   	OWF_Key[436,9]:=1170757502;
   	OWF_Key[436,10]:=379063934;
   	OWF_Key[436,11]:=939425324;
   	OWF_Key[436,12]:=1571077433;
   	OWF_Key[436,13]:=386926956;
   	OWF_Key[436,14]:=1253683460;
   	OWF_Key[436,15]:=1978140769;
   	OWF_Key[436,16]:=969971513;
   	OWF_Key[437,0]:=1843141582;
   	OWF_Key[437,1]:=1139180362;
   	OWF_Key[437,2]:=1967511731;
   	OWF_Key[437,3]:=1290649002;
   	OWF_Key[437,4]:=1378760868;
   	OWF_Key[437,5]:=1424739908;
   	OWF_Key[437,6]:=88097231;
   	OWF_Key[437,7]:=835055186;
   	OWF_Key[437,8]:=1627536833;
   	OWF_Key[437,9]:=543176006;
   	OWF_Key[437,10]:=1462679088;
   	OWF_Key[437,11]:=893832072;
   	OWF_Key[437,12]:=149893027;
   	OWF_Key[437,13]:=919941861;
   	OWF_Key[437,14]:=1244070675;
   	OWF_Key[437,15]:=720720483;
   	OWF_Key[437,16]:=106207793;
   	OWF_Key[438,0]:=1266683906;
   	OWF_Key[438,1]:=1923048867;
   	OWF_Key[438,2]:=1845235682;
   	OWF_Key[438,3]:=1052576015;
   	OWF_Key[438,4]:=621819626;
   	OWF_Key[438,5]:=249692926;
   	OWF_Key[438,6]:=969832967;
   	OWF_Key[438,7]:=766223670;
   	OWF_Key[438,8]:=1411344155;
   	OWF_Key[438,9]:=1650208802;
   	OWF_Key[438,10]:=103954679;
   	OWF_Key[438,11]:=1231682890;
   	OWF_Key[438,12]:=1324790258;
   	OWF_Key[438,13]:=615786523;
   	OWF_Key[438,14]:=414858455;
   	OWF_Key[438,15]:=939305588;
   	OWF_Key[438,16]:=719104723;
   	OWF_Key[439,0]:=1992499359;
   	OWF_Key[439,1]:=251323729;
   	OWF_Key[439,2]:=600659015;
   	OWF_Key[439,3]:=1403077275;
   	OWF_Key[439,4]:=628364857;
   	OWF_Key[439,5]:=1823764687;
   	OWF_Key[439,6]:=631857018;
   	OWF_Key[439,7]:=1931716673;
   	OWF_Key[439,8]:=428827108;
   	OWF_Key[439,9]:=1029064288;
   	OWF_Key[439,10]:=1492699981;
   	OWF_Key[439,11]:=611446466;
   	OWF_Key[439,12]:=289686517;
   	OWF_Key[439,13]:=1524542361;
   	OWF_Key[439,14]:=69099460;
   	OWF_Key[439,15]:=1294673003;
   	OWF_Key[439,16]:=2029874974;
   	OWF_Key[440,0]:=267240957;
   	OWF_Key[440,1]:=1397447859;
   	OWF_Key[440,2]:=766044100;
   	OWF_Key[440,3]:=1128726900;
   	OWF_Key[440,4]:=808363166;
   	OWF_Key[440,5]:=1558535267;
   	OWF_Key[440,6]:=1447582414;
   	OWF_Key[440,7]:=964974356;
   	OWF_Key[440,8]:=1784322886;
   	OWF_Key[440,9]:=443035495;
   	OWF_Key[440,10]:=820593840;
   	OWF_Key[440,11]:=1887778601;
   	OWF_Key[440,12]:=501962005;
   	OWF_Key[440,13]:=813962242;
   	OWF_Key[440,14]:=424069181;
   	OWF_Key[440,15]:=2011873949;
   	OWF_Key[440,16]:=1151398729;
   	OWF_Key[441,0]:=1505451756;
   	OWF_Key[441,1]:=1240333609;
   	OWF_Key[441,2]:=2098390839;
   	OWF_Key[441,3]:=1534363580;
   	OWF_Key[441,4]:=1328251268;
   	OWF_Key[441,5]:=675353205;
   	OWF_Key[441,6]:=815352173;
   	OWF_Key[441,7]:=677956491;
   	OWF_Key[441,8]:=1937060640;
   	OWF_Key[441,9]:=1410181306;
   	OWF_Key[441,10]:=758251906;
   	OWF_Key[441,11]:=1347373853;
   	OWF_Key[441,12]:=1255507361;
   	OWF_Key[441,13]:=1881254403;
   	OWF_Key[441,14]:=234983717;
   	OWF_Key[441,15]:=1703206761;
   	OWF_Key[441,16]:=1202714744;
   	OWF_Key[442,0]:=409398206;
   	OWF_Key[442,1]:=2039732025;
   	OWF_Key[442,2]:=1499250842;
   	OWF_Key[442,3]:=2021339656;
   	OWF_Key[442,4]:=1523916267;
   	OWF_Key[442,5]:=43891699;
   	OWF_Key[442,6]:=849098139;
   	OWF_Key[442,7]:=1496998499;
   	OWF_Key[442,8]:=1231230248;
   	OWF_Key[442,9]:=1160567614;
   	OWF_Key[442,10]:=1917660319;
   	OWF_Key[442,11]:=1120014121;
   	OWF_Key[442,12]:=503461202;
   	OWF_Key[442,13]:=431761410;
   	OWF_Key[442,14]:=478061027;
   	OWF_Key[442,15]:=2018840416;
   	OWF_Key[442,16]:=1866662703;
   	OWF_Key[443,0]:=1307750086;
   	OWF_Key[443,1]:=588336084;
   	OWF_Key[443,2]:=37098424;
   	OWF_Key[443,3]:=549767259;
   	OWF_Key[443,4]:=726715554;
   	OWF_Key[443,5]:=595045509;
   	OWF_Key[443,6]:=2005314031;
   	OWF_Key[443,7]:=1138018449;
   	OWF_Key[443,8]:=87073158;
   	OWF_Key[443,9]:=1057416230;
   	OWF_Key[443,10]:=1174872821;
   	OWF_Key[443,11]:=724059004;
   	OWF_Key[443,12]:=440554247;
   	OWF_Key[443,13]:=564587306;
   	OWF_Key[443,14]:=933235057;
   	OWF_Key[443,15]:=514553885;
   	OWF_Key[443,16]:=783957354;
   	OWF_Key[444,0]:=1937470562;
   	OWF_Key[444,1]:=1634266430;
   	OWF_Key[444,2]:=1078299281;
   	OWF_Key[444,3]:=2062725520;
   	OWF_Key[444,4]:=1546936069;
   	OWF_Key[444,5]:=361132692;
   	OWF_Key[444,6]:=1035953212;
   	OWF_Key[444,7]:=1703706874;
   	OWF_Key[444,8]:=1827220084;
   	OWF_Key[444,9]:=384500317;
   	OWF_Key[444,10]:=858111795;
   	OWF_Key[444,11]:=126754950;
   	OWF_Key[444,12]:=548020974;
   	OWF_Key[444,13]:=1526552867;
   	OWF_Key[444,14]:=500706782;
   	OWF_Key[444,15]:=457271281;
   	OWF_Key[444,16]:=1298806591;
   	OWF_Key[445,0]:=1152454734;
   	OWF_Key[445,1]:=1522843954;
   	OWF_Key[445,2]:=1104045148;
   	OWF_Key[445,3]:=1646359978;
   	OWF_Key[445,4]:=1910893345;
   	OWF_Key[445,5]:=275094290;
   	OWF_Key[445,6]:=490694853;
   	OWF_Key[445,7]:=1661112942;
   	OWF_Key[445,8]:=504704284;
   	OWF_Key[445,9]:=1306146160;
   	OWF_Key[445,10]:=323686031;
   	OWF_Key[445,11]:=1964751122;
   	OWF_Key[445,12]:=2076379137;
   	OWF_Key[445,13]:=1547739221;
   	OWF_Key[445,14]:=1914931196;
   	OWF_Key[445,15]:=599145780;
   	OWF_Key[445,16]:=819353237;
   	OWF_Key[446,0]:=1129528852;
   	OWF_Key[446,1]:=1855692816;
   	OWF_Key[446,2]:=1723307724;
   	OWF_Key[446,3]:=561491111;
   	OWF_Key[446,4]:=1923728612;
   	OWF_Key[446,5]:=614121178;
   	OWF_Key[446,6]:=1713617777;
   	OWF_Key[446,7]:=1457802104;
   	OWF_Key[446,8]:=516535642;
   	OWF_Key[446,9]:=535470;
   	OWF_Key[446,10]:=2048441556;
   	OWF_Key[446,11]:=2069329706;
   	OWF_Key[446,12]:=1404004704;
   	OWF_Key[446,13]:=786218775;
   	OWF_Key[446,14]:=769300157;
   	OWF_Key[446,15]:=69216967;
   	OWF_Key[446,16]:=1061177738;
   	OWF_Key[447,0]:=1467926324;
   	OWF_Key[447,1]:=1408602900;
   	OWF_Key[447,2]:=876103482;
   	OWF_Key[447,3]:=393340229;
   	OWF_Key[447,4]:=1221354422;
   	OWF_Key[447,5]:=1269305273;
   	OWF_Key[447,6]:=373849962;
   	OWF_Key[447,7]:=1887264564;
   	OWF_Key[447,8]:=1621494280;
   	OWF_Key[447,9]:=64822401;
   	OWF_Key[447,10]:=1306746888;
   	OWF_Key[447,11]:=14685194;
   	OWF_Key[447,12]:=891224843;
   	OWF_Key[447,13]:=2096386470;
   	OWF_Key[447,14]:=710798920;
   	OWF_Key[447,15]:=1361366541;
   	OWF_Key[447,16]:=628165100;
   	OWF_Key[448,0]:=1227582932;
   	OWF_Key[448,1]:=2146244073;
   	OWF_Key[448,2]:=1035592767;
   	OWF_Key[448,3]:=1797577282;
   	OWF_Key[448,4]:=983285620;
   	OWF_Key[448,5]:=1838420811;
   	OWF_Key[448,6]:=661957544;
   	OWF_Key[448,7]:=1490235311;
   	OWF_Key[448,8]:=1623052843;
   	OWF_Key[448,9]:=1831503145;
   	OWF_Key[448,10]:=1728993382;
   	OWF_Key[448,11]:=892500672;
   	OWF_Key[448,12]:=228235716;
   	OWF_Key[448,13]:=1009449319;
   	OWF_Key[448,14]:=1244627896;
   	OWF_Key[448,15]:=975416352;
   	OWF_Key[448,16]:=933233698;
   	OWF_Key[449,0]:=353168346;
   	OWF_Key[449,1]:=1990192589;
   	OWF_Key[449,2]:=1563287769;
   	OWF_Key[449,3]:=629147909;
   	OWF_Key[449,4]:=368877615;
   	OWF_Key[449,5]:=632802304;
   	OWF_Key[449,6]:=1404395808;
   	OWF_Key[449,7]:=234933487;
   	OWF_Key[449,8]:=2035753874;
   	OWF_Key[449,9]:=81487530;
   	OWF_Key[449,10]:=689508137;
   	OWF_Key[449,11]:=621812509;
   	OWF_Key[449,12]:=1127174421;
   	OWF_Key[449,13]:=232651311;
   	OWF_Key[449,14]:=1530647385;
   	OWF_Key[449,15]:=1449843934;
   	OWF_Key[449,16]:=1448221176;
   	OWF_Key[450,0]:=1480720020;
   	OWF_Key[450,1]:=971229881;
   	OWF_Key[450,2]:=39274639;
   	OWF_Key[450,3]:=2036943518;
   	OWF_Key[450,4]:=1823405599;
   	OWF_Key[450,5]:=1908461912;
   	OWF_Key[450,6]:=1869320412;
   	OWF_Key[450,7]:=578149025;
   	OWF_Key[450,8]:=1825311691;
   	OWF_Key[450,9]:=817807154;
   	OWF_Key[450,10]:=1013377412;
   	OWF_Key[450,11]:=144132748;
   	OWF_Key[450,12]:=328569765;
   	OWF_Key[450,13]:=2123802922;
   	OWF_Key[450,14]:=793248458;
   	OWF_Key[450,15]:=1267352952;
   	OWF_Key[450,16]:=1615922031;
   	OWF_Key[451,0]:=768626777;
   	OWF_Key[451,1]:=766871668;
   	OWF_Key[451,2]:=1183312167;
   	OWF_Key[451,3]:=1581685848;
   	OWF_Key[451,4]:=1708624541;
   	OWF_Key[451,5]:=786969279;
   	OWF_Key[451,6]:=1960367327;
   	OWF_Key[451,7]:=826835405;
   	OWF_Key[451,8]:=179226169;
   	OWF_Key[451,9]:=274175293;
   	OWF_Key[451,10]:=1107266177;
   	OWF_Key[451,11]:=2030652548;
   	OWF_Key[451,12]:=883467139;
   	OWF_Key[451,13]:=636829396;
   	OWF_Key[451,14]:=592001807;
   	OWF_Key[451,15]:=571497416;
   	OWF_Key[451,16]:=1868798255;
   	OWF_Key[452,0]:=516991822;
   	OWF_Key[452,1]:=207163124;
   	OWF_Key[452,2]:=59036676;
   	OWF_Key[452,3]:=1615041867;
   	OWF_Key[452,4]:=567683899;
   	OWF_Key[452,5]:=142029912;
   	OWF_Key[452,6]:=931217865;
   	OWF_Key[452,7]:=1667996348;
   	OWF_Key[452,8]:=96192727;
   	OWF_Key[452,9]:=1868114449;
   	OWF_Key[452,10]:=1301457533;
   	OWF_Key[452,11]:=286979570;
   	OWF_Key[452,12]:=880659069;
   	OWF_Key[452,13]:=577537532;
   	OWF_Key[452,14]:=153952541;
   	OWF_Key[452,15]:=1040427805;
   	OWF_Key[452,16]:=1422323838;
   	OWF_Key[453,0]:=435964332;
   	OWF_Key[453,1]:=1113581113;
   	OWF_Key[453,2]:=1037955806;
   	OWF_Key[453,3]:=832349380;
   	OWF_Key[453,4]:=1045960472;
   	OWF_Key[453,5]:=1341544677;
   	OWF_Key[453,6]:=1832789608;
   	OWF_Key[453,7]:=1578453728;
   	OWF_Key[453,8]:=26617147;
   	OWF_Key[453,9]:=696723165;
   	OWF_Key[453,10]:=987332665;
   	OWF_Key[453,11]:=2117790715;
   	OWF_Key[453,12]:=67763764;
   	OWF_Key[453,13]:=179335245;
   	OWF_Key[453,14]:=2033221386;
   	OWF_Key[453,15]:=964080003;
   	OWF_Key[453,16]:=2071944913;
   	OWF_Key[454,0]:=1112645342;
   	OWF_Key[454,1]:=1299153531;
   	OWF_Key[454,2]:=680230370;
   	OWF_Key[454,3]:=1774239879;
   	OWF_Key[454,4]:=1456417461;
   	OWF_Key[454,5]:=2028561879;
   	OWF_Key[454,6]:=1230769268;
   	OWF_Key[454,7]:=1474313834;
   	OWF_Key[454,8]:=1469609727;
   	OWF_Key[454,9]:=90773141;
   	OWF_Key[454,10]:=2137610909;
   	OWF_Key[454,11]:=919088219;
   	OWF_Key[454,12]:=308895211;
   	OWF_Key[454,13]:=1223720026;
   	OWF_Key[454,14]:=1472451160;
   	OWF_Key[454,15]:=2057853176;
   	OWF_Key[454,16]:=627927214;
   	OWF_Key[455,0]:=539678737;
   	OWF_Key[455,1]:=1496164946;
   	OWF_Key[455,2]:=1390981119;
   	OWF_Key[455,3]:=7797426;
   	OWF_Key[455,4]:=1566580114;
   	OWF_Key[455,5]:=1416421634;
   	OWF_Key[455,6]:=1098937770;
   	OWF_Key[455,7]:=2123919710;
   	OWF_Key[455,8]:=467317316;
   	OWF_Key[455,9]:=908316865;
   	OWF_Key[455,10]:=1643382700;
   	OWF_Key[455,11]:=1007088734;
   	OWF_Key[455,12]:=1350086116;
   	OWF_Key[455,13]:=269343793;
   	OWF_Key[455,14]:=1816064728;
   	OWF_Key[455,15]:=2019849996;
   	OWF_Key[455,16]:=973095462;
   	OWF_Key[456,0]:=651778823;
   	OWF_Key[456,1]:=796139351;
   	OWF_Key[456,2]:=1639774348;
   	OWF_Key[456,3]:=426142391;
   	OWF_Key[456,4]:=1510350899;
   	OWF_Key[456,5]:=1274911782;
   	OWF_Key[456,6]:=828274644;
   	OWF_Key[456,7]:=2138151514;
   	OWF_Key[456,8]:=1941572533;
   	OWF_Key[456,9]:=1637726725;
   	OWF_Key[456,10]:=1851856706;
   	OWF_Key[456,11]:=31466403;
   	OWF_Key[456,12]:=674113331;
   	OWF_Key[456,13]:=182269368;
   	OWF_Key[456,14]:=164755195;
   	OWF_Key[456,15]:=1246182194;
   	OWF_Key[456,16]:=1079651431;
   	OWF_Key[457,0]:=1338313336;
   	OWF_Key[457,1]:=1963330994;
   	OWF_Key[457,2]:=1031209559;
   	OWF_Key[457,3]:=1812457210;
   	OWF_Key[457,4]:=14121706;
   	OWF_Key[457,5]:=162931894;
   	OWF_Key[457,6]:=654115803;
   	OWF_Key[457,7]:=227249452;
   	OWF_Key[457,8]:=1934326487;
   	OWF_Key[457,9]:=349031195;
   	OWF_Key[457,10]:=86809695;
   	OWF_Key[457,11]:=1381172587;
   	OWF_Key[457,12]:=2067368640;
   	OWF_Key[457,13]:=2107491437;
   	OWF_Key[457,14]:=2072249296;
   	OWF_Key[457,15]:=669677001;
   	OWF_Key[457,16]:=37225262;
   	OWF_Key[458,0]:=1503908978;
   	OWF_Key[458,1]:=1391013770;
   	OWF_Key[458,2]:=1308639285;
   	OWF_Key[458,3]:=329039392;
   	OWF_Key[458,4]:=67714649;
   	OWF_Key[458,5]:=1749607891;
   	OWF_Key[458,6]:=1009009953;
   	OWF_Key[458,7]:=589613938;
   	OWF_Key[458,8]:=930851832;
   	OWF_Key[458,9]:=947828478;
   	OWF_Key[458,10]:=1011680299;
   	OWF_Key[458,11]:=472184037;
   	OWF_Key[458,12]:=627894634;
   	OWF_Key[458,13]:=236016349;
   	OWF_Key[458,14]:=676134881;
   	OWF_Key[458,15]:=263301723;
   	OWF_Key[458,16]:=1628619254;
   	OWF_Key[459,0]:=166177433;
   	OWF_Key[459,1]:=1589428569;
   	OWF_Key[459,2]:=607724941;
   	OWF_Key[459,3]:=280895573;
   	OWF_Key[459,4]:=1035331916;
   	OWF_Key[459,5]:=1841575505;
   	OWF_Key[459,6]:=2035399886;
   	OWF_Key[459,7]:=497272875;
   	OWF_Key[459,8]:=1342928221;
   	OWF_Key[459,9]:=357970921;
   	OWF_Key[459,10]:=328742689;
   	OWF_Key[459,11]:=682821884;
   	OWF_Key[459,12]:=1553212569;
   	OWF_Key[459,13]:=1556204228;
   	OWF_Key[459,14]:=1601258597;
   	OWF_Key[459,15]:=1356135620;
   	OWF_Key[459,16]:=811754377;
   	OWF_Key[460,0]:=1237279547;
   	OWF_Key[460,1]:=138802366;
   	OWF_Key[460,2]:=1562584751;
   	OWF_Key[460,3]:=500407363;
   	OWF_Key[460,4]:=1046562175;
   	OWF_Key[460,5]:=414710546;
   	OWF_Key[460,6]:=397688114;
   	OWF_Key[460,7]:=202760260;
   	OWF_Key[460,8]:=2141681349;
   	OWF_Key[460,9]:=1066182692;
   	OWF_Key[460,10]:=675090097;
   	OWF_Key[460,11]:=1327195608;
   	OWF_Key[460,12]:=1230339864;
   	OWF_Key[460,13]:=1662252637;
   	OWF_Key[460,14]:=2046284003;
   	OWF_Key[460,15]:=812207371;
   	OWF_Key[460,16]:=1058051825;
   	OWF_Key[461,0]:=495217914;
   	OWF_Key[461,1]:=1410369287;
   	OWF_Key[461,2]:=1705183015;
   	OWF_Key[461,3]:=1676366393;
   	OWF_Key[461,4]:=1510755823;
   	OWF_Key[461,5]:=69133510;
   	OWF_Key[461,6]:=898080451;
   	OWF_Key[461,7]:=1982025798;
   	OWF_Key[461,8]:=754232989;
   	OWF_Key[461,9]:=1425963569;
   	OWF_Key[461,10]:=774713689;
   	OWF_Key[461,11]:=895124740;
   	OWF_Key[461,12]:=1725100255;
   	OWF_Key[461,13]:=1160104106;
   	OWF_Key[461,14]:=1795787790;
   	OWF_Key[461,15]:=510470442;
   	OWF_Key[461,16]:=728898902;
   	OWF_Key[462,0]:=797747579;
   	OWF_Key[462,1]:=1942244591;
   	OWF_Key[462,2]:=1473555713;
   	OWF_Key[462,3]:=1740467233;
   	OWF_Key[462,4]:=748594188;
   	OWF_Key[462,5]:=1835855514;
   	OWF_Key[462,6]:=576453925;
   	OWF_Key[462,7]:=288875;
   	OWF_Key[462,8]:=1429835582;
   	OWF_Key[462,9]:=1556220982;
   	OWF_Key[462,10]:=1701129401;
   	OWF_Key[462,11]:=582449102;
   	OWF_Key[462,12]:=802827637;
   	OWF_Key[462,13]:=1649448373;
   	OWF_Key[462,14]:=1750880931;
   	OWF_Key[462,15]:=54162008;
   	OWF_Key[462,16]:=851938218;
   	OWF_Key[463,0]:=865670750;
   	OWF_Key[463,1]:=594716065;
   	OWF_Key[463,2]:=2034089253;
   	OWF_Key[463,3]:=2145960135;
   	OWF_Key[463,4]:=1982100569;
   	OWF_Key[463,5]:=294545367;
   	OWF_Key[463,6]:=919323143;
   	OWF_Key[463,7]:=812106562;
   	OWF_Key[463,8]:=417542431;
   	OWF_Key[463,9]:=1921837933;
   	OWF_Key[463,10]:=207393778;
   	OWF_Key[463,11]:=867003910;
   	OWF_Key[463,12]:=1734661474;
   	OWF_Key[463,13]:=415485744;
   	OWF_Key[463,14]:=1118712251;
   	OWF_Key[463,15]:=2143519391;
   	OWF_Key[463,16]:=1119215818;
   	OWF_Key[464,0]:=1737624523;
   	OWF_Key[464,1]:=1460081831;
   	OWF_Key[464,2]:=845504974;
   	OWF_Key[464,3]:=1285889610;
   	OWF_Key[464,4]:=619275188;
   	OWF_Key[464,5]:=1626633691;
   	OWF_Key[464,6]:=48888577;
   	OWF_Key[464,7]:=499455727;
   	OWF_Key[464,8]:=1108822909;
   	OWF_Key[464,9]:=649694657;
   	OWF_Key[464,10]:=1854027105;
   	OWF_Key[464,11]:=563571533;
   	OWF_Key[464,12]:=1521682057;
   	OWF_Key[464,13]:=1724655381;
   	OWF_Key[464,14]:=2051092530;
   	OWF_Key[464,15]:=645295652;
   	OWF_Key[464,16]:=442822325;
   	OWF_Key[465,0]:=276025028;
   	OWF_Key[465,1]:=538026301;
   	OWF_Key[465,2]:=475915598;
   	OWF_Key[465,3]:=180625568;
   	OWF_Key[465,4]:=389465560;
   	OWF_Key[465,5]:=1972532277;
   	OWF_Key[465,6]:=1707014637;
   	OWF_Key[465,7]:=1304612082;
   	OWF_Key[465,8]:=1408688259;
   	OWF_Key[465,9]:=1957848533;
   	OWF_Key[465,10]:=915159620;
   	OWF_Key[465,11]:=766750606;
   	OWF_Key[465,12]:=478228545;
   	OWF_Key[465,13]:=1740421605;
   	OWF_Key[465,14]:=2137954118;
   	OWF_Key[465,15]:=1217651257;
   	OWF_Key[465,16]:=965488440;
   	OWF_Key[466,0]:=979093082;
   	OWF_Key[466,1]:=1090418671;
   	OWF_Key[466,2]:=730976138;
   	OWF_Key[466,3]:=372798398;
   	OWF_Key[466,4]:=1339155871;
   	OWF_Key[466,5]:=2036204906;
   	OWF_Key[466,6]:=1287198307;
   	OWF_Key[466,7]:=1353099750;
   	OWF_Key[466,8]:=769259236;
   	OWF_Key[466,9]:=583436074;
   	OWF_Key[466,10]:=774665737;
   	OWF_Key[466,11]:=2094465580;
   	OWF_Key[466,12]:=1724883739;
   	OWF_Key[466,13]:=609152788;
   	OWF_Key[466,14]:=157706009;
   	OWF_Key[466,15]:=1044674527;
   	OWF_Key[466,16]:=1436382031;
   	OWF_Key[467,0]:=1147857297;
   	OWF_Key[467,1]:=1322618478;
   	OWF_Key[467,2]:=1887686257;
   	OWF_Key[467,3]:=2106809596;
   	OWF_Key[467,4]:=576321963;
   	OWF_Key[467,5]:=2138876048;
   	OWF_Key[467,6]:=1261440994;
   	OWF_Key[467,7]:=455915827;
   	OWF_Key[467,8]:=456592452;
   	OWF_Key[467,9]:=126113309;
   	OWF_Key[467,10]:=1033920759;
   	OWF_Key[467,11]:=1173566478;
   	OWF_Key[467,12]:=159313938;
   	OWF_Key[467,13]:=1970440684;
   	OWF_Key[467,14]:=239464061;
   	OWF_Key[467,15]:=874718528;
   	OWF_Key[467,16]:=2018261763;
   	OWF_Key[468,0]:=2016476973;
   	OWF_Key[468,1]:=92393353;
   	OWF_Key[468,2]:=994618693;
   	OWF_Key[468,3]:=1511284313;
   	OWF_Key[468,4]:=1186108722;
   	OWF_Key[468,5]:=371697827;
   	OWF_Key[468,6]:=1559784828;
   	OWF_Key[468,7]:=358433973;
   	OWF_Key[468,8]:=860249121;
   	OWF_Key[468,9]:=1328611019;
   	OWF_Key[468,10]:=1409668126;
   	OWF_Key[468,11]:=1974711422;
   	OWF_Key[468,12]:=651729088;
   	OWF_Key[468,13]:=1662744558;
   	OWF_Key[468,14]:=344073694;
   	OWF_Key[468,15]:=731530374;
   	OWF_Key[468,16]:=190518977;
   	OWF_Key[469,0]:=1691271936;
   	OWF_Key[469,1]:=1318701646;
   	OWF_Key[469,2]:=763870310;
   	OWF_Key[469,3]:=136755475;
   	OWF_Key[469,4]:=558656650;
   	OWF_Key[469,5]:=564878925;
   	OWF_Key[469,6]:=660303340;
   	OWF_Key[469,7]:=2049561079;
   	OWF_Key[469,8]:=1762628397;
   	OWF_Key[469,9]:=556772279;
   	OWF_Key[469,10]:=575942354;
   	OWF_Key[469,11]:=1088647840;
   	OWF_Key[469,12]:=802886209;
   	OWF_Key[469,13]:=149682190;
   	OWF_Key[469,14]:=1540117024;
   	OWF_Key[469,15]:=1552337669;
   	OWF_Key[469,16]:=419125738;
   	OWF_Key[470,0]:=786290986;
   	OWF_Key[470,1]:=1898352606;
   	OWF_Key[470,2]:=1860631456;
   	OWF_Key[470,3]:=1252041226;
   	OWF_Key[470,4]:=1708716096;
   	OWF_Key[470,5]:=1642111068;
   	OWF_Key[470,6]:=1444631993;
   	OWF_Key[470,7]:=1197364462;
   	OWF_Key[470,8]:=1509614677;
   	OWF_Key[470,9]:=1675323253;
   	OWF_Key[470,10]:=76303900;
   	OWF_Key[470,11]:=2077624715;
   	OWF_Key[470,12]:=115607967;
   	OWF_Key[470,13]:=821741380;
   	OWF_Key[470,14]:=884973253;
   	OWF_Key[470,15]:=1373559755;
   	OWF_Key[470,16]:=1142099432;
   	OWF_Key[471,0]:=583488049;
   	OWF_Key[471,1]:=167469148;
   	OWF_Key[471,2]:=970442439;
   	OWF_Key[471,3]:=1319743066;
   	OWF_Key[471,4]:=1458168605;
   	OWF_Key[471,5]:=1725578028;
   	OWF_Key[471,6]:=1531495223;
   	OWF_Key[471,7]:=134379754;
   	OWF_Key[471,8]:=1144126882;
   	OWF_Key[471,9]:=1296963522;
   	OWF_Key[471,10]:=1031445679;
   	OWF_Key[471,11]:=891833596;
   	OWF_Key[471,12]:=697353808;
   	OWF_Key[471,13]:=285827242;
   	OWF_Key[471,14]:=1319530;
   	OWF_Key[471,15]:=673169862;
   	OWF_Key[471,16]:=912024389;
   	OWF_Key[472,0]:=7302635;
   	OWF_Key[472,1]:=1146025357;
   	OWF_Key[472,2]:=1022331280;
   	OWF_Key[472,3]:=1729395937;
   	OWF_Key[472,4]:=791291632;
   	OWF_Key[472,5]:=313830235;
   	OWF_Key[472,6]:=954403739;
   	OWF_Key[472,7]:=630716563;
   	OWF_Key[472,8]:=1525861001;
   	OWF_Key[472,9]:=1773884953;
   	OWF_Key[472,10]:=838266152;
   	OWF_Key[472,11]:=1965223310;
   	OWF_Key[472,12]:=1724593838;
   	OWF_Key[472,13]:=1080039488;
   	OWF_Key[472,14]:=1929687523;
   	OWF_Key[472,15]:=1114222042;
   	OWF_Key[472,16]:=583718236;
   	OWF_Key[473,0]:=245279261;
   	OWF_Key[473,1]:=1371173047;
   	OWF_Key[473,2]:=468766201;
   	OWF_Key[473,3]:=990111697;
   	OWF_Key[473,4]:=76736988;
   	OWF_Key[473,5]:=1808199976;
   	OWF_Key[473,6]:=970381060;
   	OWF_Key[473,7]:=1259144862;
   	OWF_Key[473,8]:=2127722503;
   	OWF_Key[473,9]:=2091376392;
   	OWF_Key[473,10]:=1711335564;
   	OWF_Key[473,11]:=145332901;
   	OWF_Key[473,12]:=436803036;
   	OWF_Key[473,13]:=1277172253;
   	OWF_Key[473,14]:=275273133;
   	OWF_Key[473,15]:=189486762;
   	OWF_Key[473,16]:=175460621;
   	OWF_Key[474,0]:=22931542;
   	OWF_Key[474,1]:=1537077824;
   	OWF_Key[474,2]:=2066545908;
   	OWF_Key[474,3]:=1731647403;
   	OWF_Key[474,4]:=1560553187;
   	OWF_Key[474,5]:=1503856464;
   	OWF_Key[474,6]:=1333848350;
   	OWF_Key[474,7]:=480723418;
   	OWF_Key[474,8]:=1087710944;
   	OWF_Key[474,9]:=283798534;
   	OWF_Key[474,10]:=474039189;
   	OWF_Key[474,11]:=999422978;
   	OWF_Key[474,12]:=150138828;
   	OWF_Key[474,13]:=818689512;
   	OWF_Key[474,14]:=714000483;
   	OWF_Key[474,15]:=533780121;
   	OWF_Key[474,16]:=149446751;
   	OWF_Key[475,0]:=1668253040;
   	OWF_Key[475,1]:=495462062;
   	OWF_Key[475,2]:=549367101;
   	OWF_Key[475,3]:=1347586431;
   	OWF_Key[475,4]:=1532900884;
   	OWF_Key[475,5]:=1132097280;
   	OWF_Key[475,6]:=407897570;
   	OWF_Key[475,7]:=406079640;
   	OWF_Key[475,8]:=489738692;
   	OWF_Key[475,9]:=1587405245;
   	OWF_Key[475,10]:=1479331132;
   	OWF_Key[475,11]:=1109797530;
   	OWF_Key[475,12]:=217314067;
   	OWF_Key[475,13]:=1599793119;
   	OWF_Key[475,14]:=1816088977;
   	OWF_Key[475,15]:=215308357;
   	OWF_Key[475,16]:=167008321;
   	OWF_Key[476,0]:=1436245985;
   	OWF_Key[476,1]:=764480555;
   	OWF_Key[476,2]:=490115295;
   	OWF_Key[476,3]:=709460083;
   	OWF_Key[476,4]:=263841861;
   	OWF_Key[476,5]:=1062140857;
   	OWF_Key[476,6]:=768411213;
   	OWF_Key[476,7]:=848586979;
   	OWF_Key[476,8]:=1800804739;
   	OWF_Key[476,9]:=1133862195;
   	OWF_Key[476,10]:=1624666115;
   	OWF_Key[476,11]:=1084702914;
   	OWF_Key[476,12]:=1347867566;
   	OWF_Key[476,13]:=750176705;
   	OWF_Key[476,14]:=221642574;
   	OWF_Key[476,15]:=318613812;
   	OWF_Key[476,16]:=1726509360;
   	OWF_Key[477,0]:=1525691625;
   	OWF_Key[477,1]:=749081189;
   	OWF_Key[477,2]:=538627488;
   	OWF_Key[477,3]:=906259458;
   	OWF_Key[477,4]:=1015161060;
   	OWF_Key[477,5]:=142592705;
   	OWF_Key[477,6]:=817729273;
   	OWF_Key[477,7]:=224706709;
   	OWF_Key[477,8]:=1899734310;
   	OWF_Key[477,9]:=1021499912;
   	OWF_Key[477,10]:=536263534;
   	OWF_Key[477,11]:=37167737;
   	OWF_Key[477,12]:=324124446;
   	OWF_Key[477,13]:=1372264576;
   	OWF_Key[477,14]:=1929270038;
   	OWF_Key[477,15]:=1558414367;
   	OWF_Key[477,16]:=1705634615;
   	OWF_Key[478,0]:=1078944932;
   	OWF_Key[478,1]:=1682394743;
   	OWF_Key[478,2]:=1765166357;
   	OWF_Key[478,3]:=312341535;
   	OWF_Key[478,4]:=1825599611;
   	OWF_Key[478,5]:=530029376;
   	OWF_Key[478,6]:=341707261;
   	OWF_Key[478,7]:=2064396720;
   	OWF_Key[478,8]:=147719307;
   	OWF_Key[478,9]:=1294257080;
   	OWF_Key[478,10]:=1670390586;
   	OWF_Key[478,11]:=699861457;
   	OWF_Key[478,12]:=1048211397;
   	OWF_Key[478,13]:=1166571696;
   	OWF_Key[478,14]:=579034163;
   	OWF_Key[478,15]:=1887134869;
   	OWF_Key[478,16]:=1082059130;
   	OWF_Key[479,0]:=1608666085;
   	OWF_Key[479,1]:=565007198;
   	OWF_Key[479,2]:=658829031;
   	OWF_Key[479,3]:=7254357;
   	OWF_Key[479,4]:=461782101;
   	OWF_Key[479,5]:=482568642;
   	OWF_Key[479,6]:=1546106434;
   	OWF_Key[479,7]:=59640665;
   	OWF_Key[479,8]:=1829122745;
   	OWF_Key[479,9]:=1150081572;
   	OWF_Key[479,10]:=1770533657;
   	OWF_Key[479,11]:=1334481588;
   	OWF_Key[479,12]:=356956866;
   	OWF_Key[479,13]:=21579949;
   	OWF_Key[479,14]:=1508645582;
   	OWF_Key[479,15]:=1620681988;
   	OWF_Key[479,16]:=273542650;
   	OWF_Key[480,0]:=1763295348;
   	OWF_Key[480,1]:=1230802222;
   	OWF_Key[480,2]:=1803898251;
   	OWF_Key[480,3]:=69916642;
   	OWF_Key[480,4]:=1074618223;
   	OWF_Key[480,5]:=1250476337;
   	OWF_Key[480,6]:=509102101;
   	OWF_Key[480,7]:=754880795;
   	OWF_Key[480,8]:=1478007280;
   	OWF_Key[480,9]:=1535190011;
   	OWF_Key[480,10]:=740724526;
   	OWF_Key[480,11]:=1947259097;
   	OWF_Key[480,12]:=1826581338;
   	OWF_Key[480,13]:=1972522082;
   	OWF_Key[480,14]:=1849660178;
   	OWF_Key[480,15]:=1227563169;
   	OWF_Key[480,16]:=389014649;
   	OWF_Key[481,0]:=1351274052;
   	OWF_Key[481,1]:=2004167571;
   	OWF_Key[481,2]:=39641822;
   	OWF_Key[481,3]:=1463882081;
   	OWF_Key[481,4]:=1351151893;
   	OWF_Key[481,5]:=533423415;
   	OWF_Key[481,6]:=2041872037;
   	OWF_Key[481,7]:=1642753678;
   	OWF_Key[481,8]:=897716260;
   	OWF_Key[481,9]:=1030559785;
   	OWF_Key[481,10]:=553014284;
   	OWF_Key[481,11]:=1702943740;
   	OWF_Key[481,12]:=1302243419;
   	OWF_Key[481,13]:=804235717;
   	OWF_Key[481,14]:=204488863;
   	OWF_Key[481,15]:=1189763546;
   	OWF_Key[481,16]:=1717525977;
   	OWF_Key[482,0]:=818176534;
   	OWF_Key[482,1]:=1173511817;
   	OWF_Key[482,2]:=373447532;
   	OWF_Key[482,3]:=954600093;
   	OWF_Key[482,4]:=2076050192;
   	OWF_Key[482,5]:=1997775246;
   	OWF_Key[482,6]:=1160861765;
   	OWF_Key[482,7]:=556590848;
   	OWF_Key[482,8]:=776944748;
   	OWF_Key[482,9]:=433620330;
   	OWF_Key[482,10]:=434145052;
   	OWF_Key[482,11]:=1389673380;
   	OWF_Key[482,12]:=890404880;
   	OWF_Key[482,13]:=963243591;
   	OWF_Key[482,14]:=196819318;
   	OWF_Key[482,15]:=963811943;
   	OWF_Key[482,16]:=2051485366;
   	OWF_Key[483,0]:=1247133829;
   	OWF_Key[483,1]:=1092939892;
   	OWF_Key[483,2]:=1329990287;
   	OWF_Key[483,3]:=1215121384;
   	OWF_Key[483,4]:=1164514305;
   	OWF_Key[483,5]:=136882047;
   	OWF_Key[483,6]:=1920539803;
   	OWF_Key[483,7]:=148891670;
   	OWF_Key[483,8]:=917979225;
   	OWF_Key[483,9]:=107672144;
   	OWF_Key[483,10]:=1020419676;
   	OWF_Key[483,11]:=1825439059;
   	OWF_Key[483,12]:=286266849;
   	OWF_Key[483,13]:=1151725044;
   	OWF_Key[483,14]:=662830021;
   	OWF_Key[483,15]:=211930016;
   	OWF_Key[483,16]:=1365620748;
   	OWF_Key[484,0]:=1736273248;
   	OWF_Key[484,1]:=1749094378;
   	OWF_Key[484,2]:=1551240742;
   	OWF_Key[484,3]:=1649584168;
   	OWF_Key[484,4]:=1635287301;
   	OWF_Key[484,5]:=1146212040;
   	OWF_Key[484,6]:=291494453;
   	OWF_Key[484,7]:=779915129;
   	OWF_Key[484,8]:=2125851440;
   	OWF_Key[484,9]:=1357301674;
   	OWF_Key[484,10]:=362634414;
   	OWF_Key[484,11]:=13178371;
   	OWF_Key[484,12]:=855085140;
   	OWF_Key[484,13]:=220424273;
   	OWF_Key[484,14]:=318810097;
   	OWF_Key[484,15]:=730550508;
   	OWF_Key[484,16]:=1730945061;
   	OWF_Key[485,0]:=180285794;
   	OWF_Key[485,1]:=1008970945;
   	OWF_Key[485,2]:=787168105;
   	OWF_Key[485,3]:=388832873;
   	OWF_Key[485,4]:=861340082;
   	OWF_Key[485,5]:=1853207524;
   	OWF_Key[485,6]:=24378705;
   	OWF_Key[485,7]:=609137240;
   	OWF_Key[485,8]:=149768174;
   	OWF_Key[485,9]:=1195602340;
   	OWF_Key[485,10]:=2119874210;
   	OWF_Key[485,11]:=87945574;
   	OWF_Key[485,12]:=1055955521;
   	OWF_Key[485,13]:=293361835;
   	OWF_Key[485,14]:=125555862;
   	OWF_Key[485,15]:=1762069637;
   	OWF_Key[485,16]:=2144915779;
   	OWF_Key[486,0]:=358735295;
   	OWF_Key[486,1]:=1414131030;
   	OWF_Key[486,2]:=328375404;
   	OWF_Key[486,3]:=476037418;
   	OWF_Key[486,4]:=1548562159;
   	OWF_Key[486,5]:=1560146335;
   	OWF_Key[486,6]:=279967341;
   	OWF_Key[486,7]:=1717852571;
   	OWF_Key[486,8]:=84696569;
   	OWF_Key[486,9]:=2112834567;
   	OWF_Key[486,10]:=1472234344;
   	OWF_Key[486,11]:=767160443;
   	OWF_Key[486,12]:=1977809840;
   	OWF_Key[486,13]:=1816946468;
   	OWF_Key[486,14]:=6203784;
   	OWF_Key[486,15]:=1968638171;
   	OWF_Key[486,16]:=1302232862;
   	OWF_Key[487,0]:=940031665;
   	OWF_Key[487,1]:=226941860;
   	OWF_Key[487,2]:=1854183775;
   	OWF_Key[487,3]:=39542395;
   	OWF_Key[487,4]:=1146399440;
   	OWF_Key[487,5]:=1034693406;
   	OWF_Key[487,6]:=1887885129;
   	OWF_Key[487,7]:=1853791518;
   	OWF_Key[487,8]:=1206996016;
   	OWF_Key[487,9]:=993829746;
   	OWF_Key[487,10]:=1121831611;
   	OWF_Key[487,11]:=1221577384;
   	OWF_Key[487,12]:=1089553964;
   	OWF_Key[487,13]:=1504918054;
   	OWF_Key[487,14]:=325819661;
   	OWF_Key[487,15]:=1246389323;
   	OWF_Key[487,16]:=1366795814;
   	OWF_Key[488,0]:=1699305633;
   	OWF_Key[488,1]:=1206532233;
   	OWF_Key[488,2]:=1708034259;
   	OWF_Key[488,3]:=2116240674;
   	OWF_Key[488,4]:=1291934110;
   	OWF_Key[488,5]:=838336223;
   	OWF_Key[488,6]:=1018392284;
   	OWF_Key[488,7]:=1257747853;
   	OWF_Key[488,8]:=741089578;
   	OWF_Key[488,9]:=1211149795;
   	OWF_Key[488,10]:=463802342;
   	OWF_Key[488,11]:=1370237821;
   	OWF_Key[488,12]:=978763132;
   	OWF_Key[488,13]:=419151161;
   	OWF_Key[488,14]:=2135795578;
   	OWF_Key[488,15]:=1417929383;
   	OWF_Key[488,16]:=365777105;
   	OWF_Key[489,0]:=1759825414;
   	OWF_Key[489,1]:=857509565;
   	OWF_Key[489,2]:=714663553;
   	OWF_Key[489,3]:=885304376;
   	OWF_Key[489,4]:=211304816;
   	OWF_Key[489,5]:=208919928;
   	OWF_Key[489,6]:=1184926502;
   	OWF_Key[489,7]:=1803429739;
   	OWF_Key[489,8]:=1597281228;
   	OWF_Key[489,9]:=2037293023;
   	OWF_Key[489,10]:=733732701;
   	OWF_Key[489,11]:=406184872;
   	OWF_Key[489,12]:=2077483307;
   	OWF_Key[489,13]:=1039956729;
   	OWF_Key[489,14]:=818855401;
   	OWF_Key[489,15]:=869471295;
   	OWF_Key[489,16]:=527647792;
   	OWF_Key[490,0]:=1984348797;
   	OWF_Key[490,1]:=531706235;
   	OWF_Key[490,2]:=1297656937;
   	OWF_Key[490,3]:=1890677602;
   	OWF_Key[490,4]:=1151313569;
   	OWF_Key[490,5]:=960117298;
   	OWF_Key[490,6]:=291724117;
   	OWF_Key[490,7]:=1884189406;
   	OWF_Key[490,8]:=1537923568;
   	OWF_Key[490,9]:=1183156426;
   	OWF_Key[490,10]:=2014099253;
   	OWF_Key[490,11]:=1819971836;
   	OWF_Key[490,12]:=1448526659;
   	OWF_Key[490,13]:=1737198382;
   	OWF_Key[490,14]:=1734796253;
   	OWF_Key[490,15]:=2070478395;
   	OWF_Key[490,16]:=937705773;
   	OWF_Key[491,0]:=1908366843;
   	OWF_Key[491,1]:=636980225;
   	OWF_Key[491,2]:=1322298004;
   	OWF_Key[491,3]:=323026572;
   	OWF_Key[491,4]:=1874382231;
   	OWF_Key[491,5]:=1024803106;
   	OWF_Key[491,6]:=1819865040;
   	OWF_Key[491,7]:=593661108;
   	OWF_Key[491,8]:=702483164;
   	OWF_Key[491,9]:=1492390470;
   	OWF_Key[491,10]:=446725061;
   	OWF_Key[491,11]:=733227282;
   	OWF_Key[491,12]:=537101106;
   	OWF_Key[491,13]:=1180544438;
   	OWF_Key[491,14]:=39922459;
   	OWF_Key[491,15]:=1190138631;
   	OWF_Key[491,16]:=1345075058;
   	OWF_Key[492,0]:=1334949409;
   	OWF_Key[492,1]:=1196430000;
   	OWF_Key[492,2]:=488884062;
   	OWF_Key[492,3]:=851550411;
   	OWF_Key[492,4]:=771475192;
   	OWF_Key[492,5]:=189712440;
   	OWF_Key[492,6]:=2101761244;
   	OWF_Key[492,7]:=1037132449;
   	OWF_Key[492,8]:=2098094500;
   	OWF_Key[492,9]:=2117658873;
   	OWF_Key[492,10]:=139600672;
   	OWF_Key[492,11]:=938272757;
   	OWF_Key[492,12]:=809032924;
   	OWF_Key[492,13]:=1945131536;
   	OWF_Key[492,14]:=271917884;
   	OWF_Key[492,15]:=514787145;
   	OWF_Key[492,16]:=1892040543;
   	OWF_Key[493,0]:=1176177756;
   	OWF_Key[493,1]:=1476281003;
   	OWF_Key[493,2]:=1329499056;
   	OWF_Key[493,3]:=876307819;
   	OWF_Key[493,4]:=1336701859;
   	OWF_Key[493,5]:=908163176;
   	OWF_Key[493,6]:=587219204;
   	OWF_Key[493,7]:=1825097095;
   	OWF_Key[493,8]:=1991583801;
   	OWF_Key[493,9]:=292409901;
   	OWF_Key[493,10]:=1655431309;
   	OWF_Key[493,11]:=1558270048;
   	OWF_Key[493,12]:=121380095;
   	OWF_Key[493,13]:=909630627;
   	OWF_Key[493,14]:=1764278601;
   	OWF_Key[493,15]:=89397778;
   	OWF_Key[493,16]:=1408732431;
   	OWF_Key[494,0]:=49553222;
   	OWF_Key[494,1]:=530494636;
   	OWF_Key[494,2]:=1284362047;
   	OWF_Key[494,3]:=311138190;
   	OWF_Key[494,4]:=1591643317;
   	OWF_Key[494,5]:=1493168117;
   	OWF_Key[494,6]:=456170775;
   	OWF_Key[494,7]:=1970021990;
   	OWF_Key[494,8]:=1169189263;
   	OWF_Key[494,9]:=680780058;
   	OWF_Key[494,10]:=893188666;
   	OWF_Key[494,11]:=990393848;
   	OWF_Key[494,12]:=1241010746;
   	OWF_Key[494,13]:=146128889;
   	OWF_Key[494,14]:=1062608701;
   	OWF_Key[494,15]:=420179203;
   	OWF_Key[494,16]:=922343458;
   	OWF_Key[495,0]:=1091769659;
   	OWF_Key[495,1]:=566809994;
   	OWF_Key[495,2]:=1077976928;
   	OWF_Key[495,3]:=1994957392;
   	OWF_Key[495,4]:=973447049;
   	OWF_Key[495,5]:=878633857;
   	OWF_Key[495,6]:=1540181116;
   	OWF_Key[495,7]:=1990232201;
   	OWF_Key[495,8]:=1526133929;
   	OWF_Key[495,9]:=2089262270;
   	OWF_Key[495,10]:=441295542;
   	OWF_Key[495,11]:=1291674150;
   	OWF_Key[495,12]:=2076895120;
   	OWF_Key[495,13]:=292865479;
   	OWF_Key[495,14]:=2074870027;
   	OWF_Key[495,15]:=2042511207;
   	OWF_Key[495,16]:=745705537;
   	OWF_Key[496,0]:=1341511840;
   	OWF_Key[496,1]:=1019466133;
   	OWF_Key[496,2]:=303481277;
   	OWF_Key[496,3]:=2007417496;
   	OWF_Key[496,4]:=1780224295;
   	OWF_Key[496,5]:=620879742;
   	OWF_Key[496,6]:=27001078;
   	OWF_Key[496,7]:=15003457;
   	OWF_Key[496,8]:=1690673941;
   	OWF_Key[496,9]:=275106391;
   	OWF_Key[496,10]:=1070017495;
   	OWF_Key[496,11]:=1530183127;
   	OWF_Key[496,12]:=2066170899;
   	OWF_Key[496,13]:=2114312374;
   	OWF_Key[496,14]:=1552826616;
   	OWF_Key[496,15]:=1214324720;
   	OWF_Key[496,16]:=775970867;
   	OWF_Key[497,0]:=111476704;
   	OWF_Key[497,1]:=120976930;
   	OWF_Key[497,2]:=673893139;
   	OWF_Key[497,3]:=1369509872;
   	OWF_Key[497,4]:=709227868;
   	OWF_Key[497,5]:=612813412;
   	OWF_Key[497,6]:=927834295;
   	OWF_Key[497,7]:=114850789;
   	OWF_Key[497,8]:=1177277687;
   	OWF_Key[497,9]:=1823004275;
   	OWF_Key[497,10]:=1000239619;
   	OWF_Key[497,11]:=327954370;
   	OWF_Key[497,12]:=54958664;
   	OWF_Key[497,13]:=825998369;
   	OWF_Key[497,14]:=473143646;
   	OWF_Key[497,15]:=1940175727;
   	OWF_Key[497,16]:=2115626236;
   	OWF_Key[498,0]:=154289919;
   	OWF_Key[498,1]:=1367598128;
   	OWF_Key[498,2]:=248930509;
   	OWF_Key[498,3]:=479332167;
   	OWF_Key[498,4]:=1430457870;
   	OWF_Key[498,5]:=319002340;
   	OWF_Key[498,6]:=1040529396;
   	OWF_Key[498,7]:=191631304;
   	OWF_Key[498,8]:=1601716912;
   	OWF_Key[498,9]:=62908199;
   	OWF_Key[498,10]:=1841559220;
   	OWF_Key[498,11]:=51252082;
   	OWF_Key[498,12]:=1844901406;
   	OWF_Key[498,13]:=789024788;
   	OWF_Key[498,14]:=1487654993;
   	OWF_Key[498,15]:=1781500674;
   	OWF_Key[498,16]:=2082739431;
   	OWF_Key[499,0]:=1507480372;
   	OWF_Key[499,1]:=570420337;
   	OWF_Key[499,2]:=15511095;
   	OWF_Key[499,3]:=2041256578;
   	OWF_Key[499,4]:=735279621;
   	OWF_Key[499,5]:=1815189437;
   	OWF_Key[499,6]:=1319098589;
   	OWF_Key[499,7]:=2057890135;
   	OWF_Key[499,8]:=305394075;
   	OWF_Key[499,9]:=1307110635;
   	OWF_Key[499,10]:=1748491928;
   	OWF_Key[499,11]:=398848138;
   	OWF_Key[499,12]:=1227950992;
   	OWF_Key[499,13]:=1565246236;
   	OWF_Key[499,14]:=533840425;
   	OWF_Key[499,15]:=25675421;
   	OWF_Key[499,16]:=1074649065;
   	OWF_Key[500,0]:=2087758853;
   	OWF_Key[500,1]:=2117589021;
   	OWF_Key[500,2]:=381542162;
   	OWF_Key[500,3]:=1738873576;
   	OWF_Key[500,4]:=1962182605;
   	OWF_Key[500,5]:=1194095748;
   	OWF_Key[500,6]:=439692198;
   	OWF_Key[500,7]:=666871853;
   	OWF_Key[500,8]:=1923530676;
   	OWF_Key[500,9]:=1040880210;
   	OWF_Key[500,10]:=356101733;
   	OWF_Key[500,11]:=1070527908;
   	OWF_Key[500,12]:=1588914785;
   	OWF_Key[500,13]:=1278126667;
   	OWF_Key[500,14]:=1673450629;
   	OWF_Key[500,15]:=1521337470;
   	OWF_Key[500,16]:=1939071007;
   	OWF_Key[501,0]:=345749202;
   	OWF_Key[501,1]:=1368887386;
   	OWF_Key[501,2]:=507225857;
   	OWF_Key[501,3]:=1763940532;
   	OWF_Key[501,4]:=1804731464;
   	OWF_Key[501,5]:=646067272;
   	OWF_Key[501,6]:=1457248766;
   	OWF_Key[501,7]:=1971973486;
   	OWF_Key[501,8]:=1353785629;
   	OWF_Key[501,9]:=2060837739;
   	OWF_Key[501,10]:=1384782142;
   	OWF_Key[501,11]:=213990247;
   	OWF_Key[501,12]:=1025391067;
   	OWF_Key[501,13]:=1924113463;
   	OWF_Key[501,14]:=1653143275;
   	OWF_Key[501,15]:=198232743;
   	OWF_Key[501,16]:=1583266005;
   	OWF_Key[502,0]:=1169360493;
   	OWF_Key[502,1]:=1136628196;
   	OWF_Key[502,2]:=366206674;
   	OWF_Key[502,3]:=297035550;
   	OWF_Key[502,4]:=573017730;
   	OWF_Key[502,5]:=1808646128;
   	OWF_Key[502,6]:=900274949;
   	OWF_Key[502,7]:=1065961152;
   	OWF_Key[502,8]:=427946820;
   	OWF_Key[502,9]:=130812029;
   	OWF_Key[502,10]:=779119194;
   	OWF_Key[502,11]:=1787344868;
   	OWF_Key[502,12]:=631265576;
   	OWF_Key[502,13]:=289088048;
   	OWF_Key[502,14]:=471820134;
   	OWF_Key[502,15]:=715034899;
   	OWF_Key[502,16]:=314698490;
   	OWF_Key[503,0]:=417246403;
   	OWF_Key[503,1]:=300717064;
   	OWF_Key[503,2]:=909286660;
   	OWF_Key[503,3]:=297352639;
   	OWF_Key[503,4]:=833884686;
   	OWF_Key[503,5]:=1135282217;
   	OWF_Key[503,6]:=676619777;
   	OWF_Key[503,7]:=221049003;
   	OWF_Key[503,8]:=1405752048;
   	OWF_Key[503,9]:=83917254;
   	OWF_Key[503,10]:=5135867;
   	OWF_Key[503,11]:=466733209;
   	OWF_Key[503,12]:=1804006315;
   	OWF_Key[503,13]:=1254553323;
   	OWF_Key[503,14]:=415869850;
   	OWF_Key[503,15]:=1883907262;
   	OWF_Key[503,16]:=1142258667;
   	OWF_Key[504,0]:=418136412;
   	OWF_Key[504,1]:=356795212;
   	OWF_Key[504,2]:=1668757104;
   	OWF_Key[504,3]:=938155562;
   	OWF_Key[504,4]:=481820915;
   	OWF_Key[504,5]:=246145341;
   	OWF_Key[504,6]:=330083365;
   	OWF_Key[504,7]:=1728047647;
   	OWF_Key[504,8]:=580062916;
   	OWF_Key[504,9]:=1726536693;
   	OWF_Key[504,10]:=1210280130;
   	OWF_Key[504,11]:=1996762682;
   	OWF_Key[504,12]:=2146543310;
   	OWF_Key[504,13]:=902315416;
   	OWF_Key[504,14]:=1682338519;
   	OWF_Key[504,15]:=1960841521;
   	OWF_Key[504,16]:=138300783;
   	OWF_Key[505,0]:=1449213295;
   	OWF_Key[505,1]:=995645721;
   	OWF_Key[505,2]:=230989164;
   	OWF_Key[505,3]:=1252878380;
   	OWF_Key[505,4]:=2105708041;
   	OWF_Key[505,5]:=483522129;
   	OWF_Key[505,6]:=704278147;
   	OWF_Key[505,7]:=2070095564;
   	OWF_Key[505,8]:=359638141;
   	OWF_Key[505,9]:=7788716;
   	OWF_Key[505,10]:=34641999;
   	OWF_Key[505,11]:=69163842;
   	OWF_Key[505,12]:=1137676405;
   	OWF_Key[505,13]:=2009012345;
   	OWF_Key[505,14]:=355914891;
   	OWF_Key[505,15]:=383472726;
   	OWF_Key[505,16]:=370509173;
   	OWF_Key[506,0]:=1887736376;
   	OWF_Key[506,1]:=1478706889;
   	OWF_Key[506,2]:=303112024;
   	OWF_Key[506,3]:=558798070;
   	OWF_Key[506,4]:=1856827029;
   	OWF_Key[506,5]:=490905567;
   	OWF_Key[506,6]:=155094389;
   	OWF_Key[506,7]:=685235939;
   	OWF_Key[506,8]:=1009793856;
   	OWF_Key[506,9]:=742817189;
   	OWF_Key[506,10]:=1616863440;
   	OWF_Key[506,11]:=907701962;
   	OWF_Key[506,12]:=1290213235;
   	OWF_Key[506,13]:=1588803444;
   	OWF_Key[506,14]:=986454397;
   	OWF_Key[506,15]:=1817296275;
   	OWF_Key[506,16]:=2131318438;
   	OWF_Key[507,0]:=1263915048;
   	OWF_Key[507,1]:=884428699;
   	OWF_Key[507,2]:=784999756;
   	OWF_Key[507,3]:=871274234;
   	OWF_Key[507,4]:=94819218;
   	OWF_Key[507,5]:=1731981740;
   	OWF_Key[507,6]:=1806819302;
   	OWF_Key[507,7]:=2032488522;
   	OWF_Key[507,8]:=1927013779;
   	OWF_Key[507,9]:=1991399524;
   	OWF_Key[507,10]:=1255862050;
   	OWF_Key[507,11]:=1975435926;
   	OWF_Key[507,12]:=2053875446;
   	OWF_Key[507,13]:=1909139500;
   	OWF_Key[507,14]:=721045760;
   	OWF_Key[507,15]:=979825626;
   	OWF_Key[507,16]:=1730626985;
   	OWF_Key[508,0]:=515328070;
   	OWF_Key[508,1]:=845401025;
   	OWF_Key[508,2]:=567423216;
   	OWF_Key[508,3]:=874781597;
   	OWF_Key[508,4]:=143310526;
   	OWF_Key[508,5]:=193648362;
   	OWF_Key[508,6]:=203250012;
   	OWF_Key[508,7]:=123594147;
   	OWF_Key[508,8]:=180272894;
   	OWF_Key[508,9]:=30188514;
   	OWF_Key[508,10]:=1656271933;
   	OWF_Key[508,11]:=752935026;
   	OWF_Key[508,12]:=1353976195;
   	OWF_Key[508,13]:=1978097901;
   	OWF_Key[508,14]:=972235183;
   	OWF_Key[508,15]:=2008401032;
   	OWF_Key[508,16]:=1196670965;
   	OWF_Key[509,0]:=1603553372;
   	OWF_Key[509,1]:=29145678;
   	OWF_Key[509,2]:=834613877;
   	OWF_Key[509,3]:=101299579;
   	OWF_Key[509,4]:=1009354627;
   	OWF_Key[509,5]:=153939168;
   	OWF_Key[509,6]:=221534287;
   	OWF_Key[509,7]:=1405378524;
   	OWF_Key[509,8]:=1891966145;
   	OWF_Key[509,9]:=668823906;
   	OWF_Key[509,10]:=1944869940;
   	OWF_Key[509,11]:=1977736820;
   	OWF_Key[509,12]:=266671220;
   	OWF_Key[509,13]:=715545849;
   	OWF_Key[509,14]:=1094288399;
   	OWF_Key[509,15]:=47243315;
   	OWF_Key[509,16]:=1532012269;
   	OWF_Key[510,0]:=1625431590;
   	OWF_Key[510,1]:=2133326443;
   	OWF_Key[510,2]:=1474462327;
   	OWF_Key[510,3]:=1740254308;
   	OWF_Key[510,4]:=911800255;
   	OWF_Key[510,5]:=405624622;
   	OWF_Key[510,6]:=2038366152;
   	OWF_Key[510,7]:=993684018;
   	OWF_Key[510,8]:=193524294;
   	OWF_Key[510,9]:=1063017460;
   	OWF_Key[510,10]:=1237814456;
   	OWF_Key[510,11]:=1258022554;
   	OWF_Key[510,12]:=1675220301;
   	OWF_Key[510,13]:=194402205;
   	OWF_Key[510,14]:=1733294351;
   	OWF_Key[510,15]:=2025100591;
   	OWF_Key[510,16]:=1557005965;
   	OWF_Key[511,0]:=1291710574;
   	OWF_Key[511,1]:=2056626527;
   	OWF_Key[511,2]:=54206082;
   	OWF_Key[511,3]:=574008565;
   	OWF_Key[511,4]:=517724135;
   	OWF_Key[511,5]:=1310685575;
   	OWF_Key[511,6]:=311040526;
   	OWF_Key[511,7]:=1632169611;
   	OWF_Key[511,8]:=1699044668;
   	OWF_Key[511,9]:=1845130475;
   	OWF_Key[511,10]:=206920097;
   	OWF_Key[511,11]:=2836175;
   	OWF_Key[511,12]:=167247896;
   	OWF_Key[511,13]:=699824645;
   	OWF_Key[511,14]:=175797739;
   	OWF_Key[511,15]:=125481641;
   	OWF_Key[511,16]:=2076761660;
   End_If;
   
END_ROUTINE
